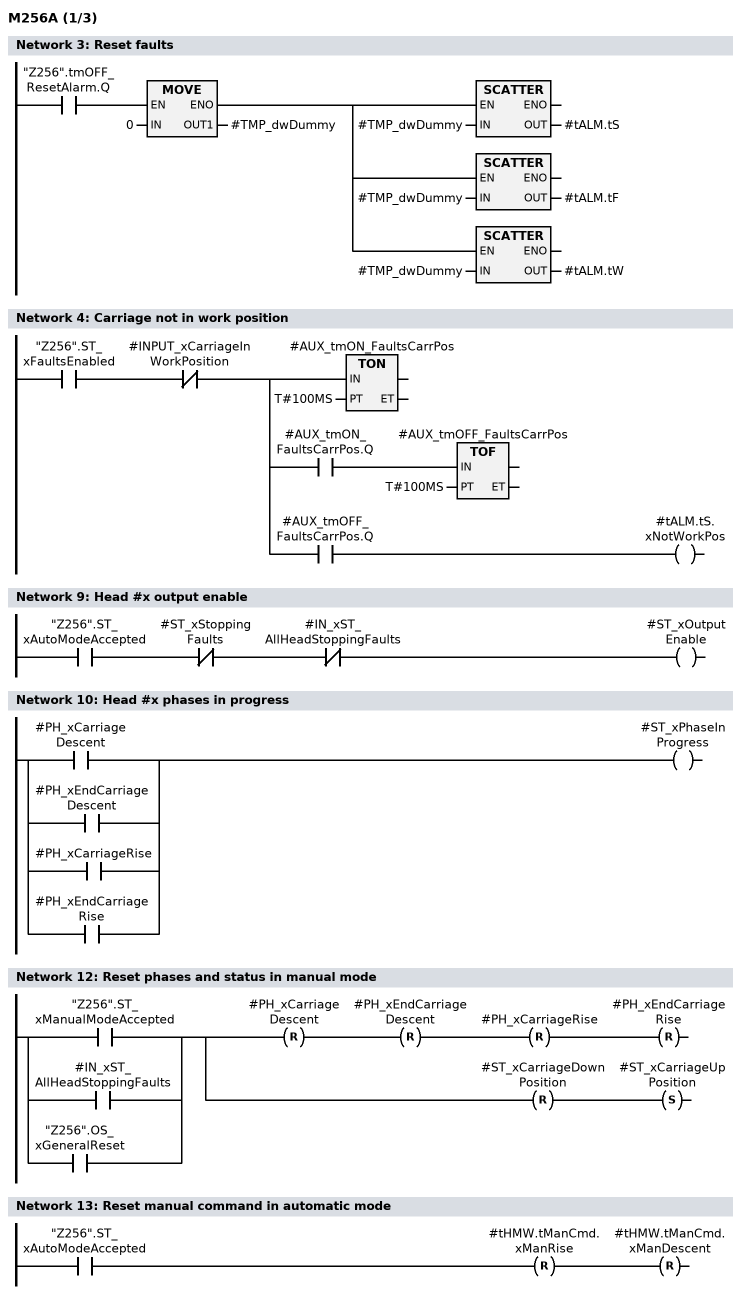
   IF "Z256".tmOFF_ResetAlarm.Q THEN #TMP_dwDummy := 0; END_IF;
   #_w1 := "Z256".tmOFF_ResetAlarm.Q;
   IF #_w1 THEN
       SCATTER(IN := #TMP_dwDummy, OUT => #tALM.tS);
       SCATTER(IN := #TMP_dwDummy, OUT => #tALM.tF);
       SCATTER(IN := #TMP_dwDummy, OUT => #tALM.tW);
   END_IF;
END_REGION

REGION Network 4: Carriage not in work position
   #_w1 := "Z256".ST_xFaultsEnabled AND NOT #INPUT_xCarriageInWorkPosition;
   #AUX_tmON_FaultsCarrPos.TON(IN := #_w1, PT := T#100MS);
   #AUX_tmOFF_FaultsCarrPos.TOF(IN := #_w1 AND #AUX_tmON_FaultsCarrPos.Q, PT := T#100MS);
   #tALM.tS.xNotWorkPos := #_w1 AND #AUX_tmOFF_FaultsCarrPos.Q;
END_REGION

REGION Network 5 (SCL): Cumulative of warning active
   #ST_xWarnings := 0;

   GATHER(IN:= #tALM.tW,
          OUT=>#TMP_dwDummy);

   IF #TMP_dwDummy <> 0 THEN
       #ST_xWarnings := 1;
   END_IF;
END_REGION

REGION Network 6 (SCL): Cumulative of stopping faults active
   #ST_xStoppingFaults := 0;
   GATHER(IN := #tALM.tS,
          OUT => #TMP_dwDummy);

   IF #TMP_dwDummy <> 0 THEN
       #ST_xStoppingFaults := 1;
   END_IF;
END_REGION

REGION Network 7 (SCL): Cumulative of faults active
   #ST_xFaults := 0;
   GATHER(IN := #tALM.tF,
          OUT => #TMP_dwDummy);

   IF #TMP_dwDummy <> 0 THEN
       #ST_xFaults := 1;
   END_IF;
END_REGION

REGION Network 8: ####_STATUS_####
END_REGION

REGION Network 9: Head #x output enable
   RUNG wire#powerrail
      Contact( "Z256".ST_xAutoModeAccepted )
      I_Contact( #ST_xStoppingFaults )
      I_Contact( #IN_xST_AllHeadStoppingFaults )
      Coil( #ST_xOutputEnable )
   END_RUNG
   // the same network as SCL:
   #ST_xOutputEnable := "Z256".ST_xAutoModeAccepted AND NOT #ST_xStoppingFaults AND NOT #IN_xST_AllHeadStoppingFaults;
END_REGION

REGION Network 10: Head #x phases in progress
   RUNG wire#powerrail
      Contact( #PH_xCarriageDescent )
      wire#w1
      Coil( #ST_xPhaseInProgress )
   END_RUNG
   RUNG wire#powerrail
      Contact( #PH_xEndCarriageDescent )
   END_RUNG wire#w1
   RUNG wire#powerrail
      Contact( #PH_xCarriageRise )
   END_RUNG wire#w1
   RUNG wire#powerrail
      Contact( #PH_xEndCarriageRise )
   END_RUNG wire#w1
   // the same network as SCL:
   #ST_xPhaseInProgress := #PH_xCarriageDescent OR #PH_xEndCarriageDescent OR #PH_xCarriageRise OR #PH_xEndCarriageRise;
END_REGION

REGION Network 11: #####_PHASES_&_LOGICS_#####
END_REGION

REGION Network 12: Reset phases and status in manual mode
   RUNG wire#powerrail
      Contact( "Z256".ST_xManualModeAccepted )
      wire#w1
      R_Coil( #PH_xCarriageDescent )
      R_Coil( #PH_xEndCarriageDescent )
      R_Coil( #PH_xCarriageRise )
      R_Coil( #PH_xEndCarriageRise )
   END_RUNG
   RUNG wire#powerrail
      Contact( #IN_xST_AllHeadStoppingFaults )
   END_RUNG wire#w1
   RUNG wire#powerrail
      Contact( "Z256".OS_xGeneralReset )
   END_RUNG wire#w1
   RUNG wire#w1
      R_Coil( #ST_xCarriageDownPosition )
      S_Coil( #ST_xCarriageUpPosition )
   END_RUNG
   // the same network as SCL:
   IF "Z256".ST_xManualModeAccepted OR #IN_xST_AllHeadStoppingFaults OR "Z256".OS_xGeneralReset THEN
       #PH_xCarriageDescent := FALSE;
       #PH_xEndCarriageDescent := FALSE;
       #PH_xCarriageRise := FALSE;
       #PH_xEndCarriageRise := FALSE;
       #ST_xCarriageDownPosition := FALSE;
       #ST_xCarriageUpPosition := TRUE;
   END_IF;
END_REGION

REGION Network 13: Reset manual command in automatic mode
   RUNG wire#powerrail
      Contact( "Z256".ST_xAutoModeAccepted )
      R_Coil( #tHMW.tManCmd.xManRise )
      R_Coil( #tHMW.tManCmd.xManDescent )
   END_RUNG
   // the same network as SCL:
   IF "Z256".ST_xAutoModeAccepted THEN
       #tHMW.tManCmd.xManRise := FALSE;
       #tHMW.tManCmd.xManDescent := FALSE;
   END_IF;
END_REGION

REGION Network 14: Carriage descent request
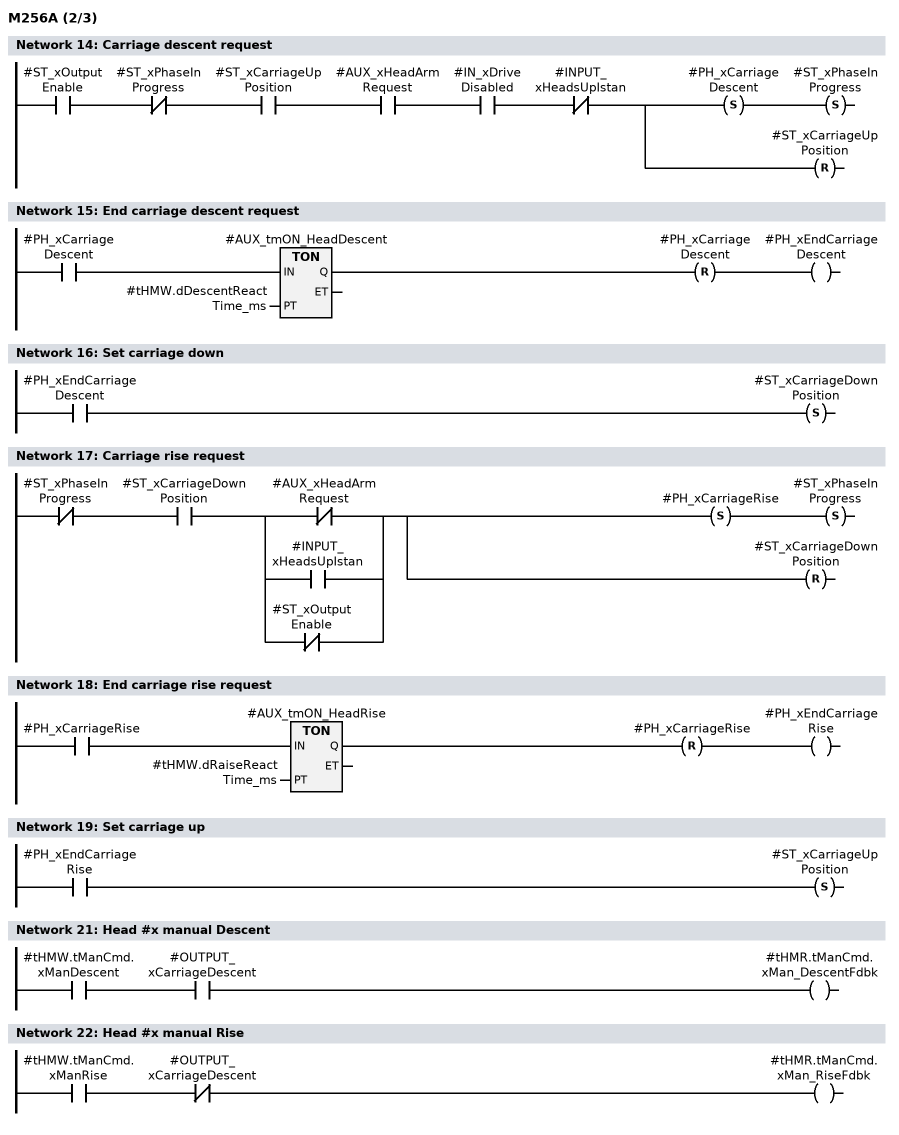
   RUNG wire#powerrail
      Contact( #ST_xOutputEnable )
      I_Contact( #ST_xPhaseInProgress )
      Contact( #ST_xCarriageUpPosition )
      Contact( #AUX_xHeadArmRequest )
      Contact( #IN_xDriveDisabled )
      I_Contact( #INPUT_xHeadsUpIstan )
      wire#w1
      S_Coil( #PH_xCarriageDescent )
      S_Coil( #ST_xPhaseInProgress )
   END_RUNG
   RUNG wire#w1
      R_Coil( #ST_xCarriageUpPosition )
   END_RUNG
   // the same network as SCL:
   IF #ST_xOutputEnable AND NOT #ST_xPhaseInProgress AND #ST_xCarriageUpPosition AND #AUX_xHeadArmRequest AND #IN_xDriveDisabled AND NOT #INPUT_xHeadsUpIstan THEN
       #PH_xCarriageDescent := TRUE;
   END_IF;
   #_w1 := #ST_xOutputEnable AND NOT #ST_xPhaseInProgress AND #ST_xCarriageUpPosition AND #AUX_xHeadArmRequest AND #IN_xDriveDisabled AND NOT #INPUT_xHeadsUpIstan;
   IF #_w1 THEN
       #ST_xPhaseInProgress := TRUE;
       #ST_xCarriageUpPosition := FALSE;
   END_IF;
END_REGION

REGION Network 15: End carriage descent request
   #AUX_tmON_HeadDescent.TON(IN := #PH_xCarriageDescent, PT := #tHMW.dDescentReactTime_ms);
   IF #AUX_tmON_HeadDescent.Q THEN #PH_xCarriageDescent := FALSE; END_IF;
   #PH_xEndCarriageDescent := #AUX_tmON_HeadDescent.Q;
END_REGION

REGION Network 16: Set carriage down
   RUNG wire#powerrail
      Contact( #PH_xEndCarriageDescent )
      S_Coil( #ST_xCarriageDownPosition )
   END_RUNG
   // the same network as SCL:
   IF #PH_xEndCarriageDescent THEN #ST_xCarriageDownPosition := TRUE; END_IF;
END_REGION

REGION Network 17: Carriage rise request
   RUNG wire#powerrail
      I_Contact( #ST_xPhaseInProgress )
      Contact( #ST_xCarriageDownPosition )
      wire#w1
      I_Contact( #AUX_xHeadArmRequest )
      wire#w2
      S_Coil( #PH_xCarriageRise )
      S_Coil( #ST_xPhaseInProgress )
   END_RUNG
   RUNG wire#w1
      Contact( #INPUT_xHeadsUpIstan )
   END_RUNG wire#w2
   RUNG wire#w1
      I_Contact( #ST_xOutputEnable )
   END_RUNG wire#w2
   RUNG wire#w2
      R_Coil( #ST_xCarriageDownPosition )
   END_RUNG
   // the same network as SCL:
   IF NOT #ST_xPhaseInProgress AND #ST_xCarriageDownPosition AND (NOT #AUX_xHeadArmRequest OR #INPUT_xHeadsUpIstan OR NOT #ST_xOutputEnable) THEN
       #PH_xCarriageRise := TRUE;
   END_IF;
   #_w1 := NOT #ST_xPhaseInProgress AND #ST_xCarriageDownPosition AND (NOT #AUX_xHeadArmRequest OR #INPUT_xHeadsUpIstan OR NOT #ST_xOutputEnable);
   IF #_w1 THEN
       #ST_xPhaseInProgress := TRUE;
       #ST_xCarriageDownPosition := FALSE;
   END_IF;
END_REGION

REGION Network 18: End carriage rise request
   #AUX_tmON_HeadRise.TON(IN := #PH_xCarriageRise, PT := #tHMW.dRaiseReactTime_ms);
   IF #AUX_tmON_HeadRise.Q THEN #PH_xCarriageRise := FALSE; END_IF;
   #PH_xEndCarriageRise := #AUX_tmON_HeadRise.Q;
END_REGION

REGION Network 19: Set carriage up
   RUNG wire#powerrail
      Contact( #PH_xEndCarriageRise )
      S_Coil( #ST_xCarriageUpPosition )
   END_RUNG
   // the same network as SCL:
   IF #PH_xEndCarriageRise THEN #ST_xCarriageUpPosition := TRUE; END_IF;
END_REGION

REGION Network 20: ### HMI STATUS ###
END_REGION

REGION Network 21: Head #x manual Descent
   RUNG wire#powerrail
      Contact( #tHMW.tManCmd.xManDescent )
      Contact( #OUTPUT_xCarriageDescent )
      Coil( #tHMR.tManCmd.xMan_DescentFdbk )
   END_RUNG
   // the same network as SCL:
   #tHMR.tManCmd.xMan_DescentFdbk := #tHMW.tManCmd.xManDescent AND #OUTPUT_xCarriageDescent;
END_REGION

REGION Network 22: Head #x manual Rise
   RUNG wire#powerrail
      Contact( #tHMW.tManCmd.xManRise )
      I_Contact( #OUTPUT_xCarriageDescent )
      Coil( #tHMR.tManCmd.xMan_RiseFdbk )
   END_RUNG
   // the same network as SCL:
   #tHMR.tManCmd.xMan_RiseFdbk := #tHMW.tManCmd.xManRise AND NOT #OUTPUT_xCarriageDescent;
END_REGION

REGION Network 23: Arm status
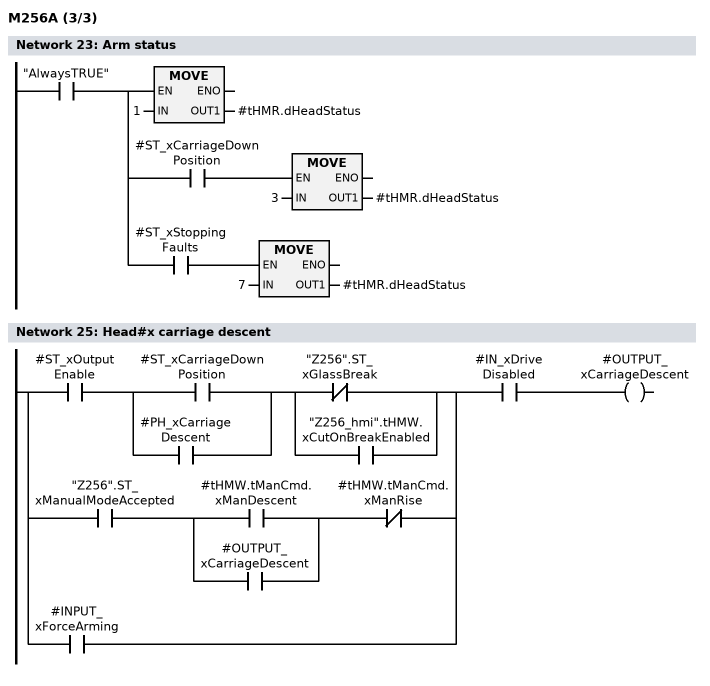
   RUNG wire#powerrail
      Contact( "AlwaysTRUE" )
      wire#w1
      Move(in := 1, out1 => #tHMR.dHeadStatus)
   END_RUNG
   RUNG wire#w1
      Contact( #ST_xCarriageDownPosition )
      Move(in := 3, out1 => #tHMR.dHeadStatus)
   END_RUNG
   RUNG wire#w1
      Contact( #ST_xStoppingFaults )
      Move(in := 7, out1 => #tHMR.dHeadStatus)
   END_RUNG
   // the same network as SCL:
   IF "AlwaysTRUE" THEN #tHMR.dHeadStatus := 1; END_IF;
   IF "AlwaysTRUE" AND #ST_xCarriageDownPosition THEN #tHMR.dHeadStatus := 3; END_IF;
   IF "AlwaysTRUE" AND #ST_xStoppingFaults THEN #tHMR.dHeadStatus := 7; END_IF;
END_REGION

REGION Network 24: ####_OUTPUT_####
END_REGION

REGION Network 25: Head#x carriage descent
   RUNG wire#powerrail
      Contact( #ST_xOutputEnable )
      wire#w1
      Contact( #ST_xCarriageDownPosition )
      wire#w2
      I_Contact( "Z256".ST_xGlassBreak )
      wire#w3
      Contact( #IN_xDriveDisabled )
      Coil( #OUTPUT_xCarriageDescent )
   END_RUNG
   RUNG wire#w1
      Contact( #PH_xCarriageDescent )
   END_RUNG wire#w2
   RUNG wire#w2
      Contact( "Z256_hmi".tHMW.xCutOnBreakEnabled )
   END_RUNG wire#w3
   RUNG wire#powerrail
      Contact( "Z256".ST_xManualModeAccepted )
      wire#w4
      Contact( #tHMW.tManCmd.xManDescent )
      wire#w5
      I_Contact( #tHMW.tManCmd.xManRise )
   END_RUNG wire#w3
   RUNG wire#w4
      Contact( #OUTPUT_xCarriageDescent )
   END_RUNG wire#w5
   RUNG wire#powerrail
      Contact( #INPUT_xForceArming )
   END_RUNG wire#w3
   // the same network as SCL:
   #OUTPUT_xCarriageDescent := ((#ST_xOutputEnable AND (#ST_xCarriageDownPosition OR #PH_xCarriageDescent) AND (NOT "Z256".ST_xGlassBreak OR "Z256_hmi".tHMW.xCutOnBreakEnabled)) OR ("Z256".ST_xManualModeAccepted AND (#tHMW.tManCmd.xManDescent OR #OUTPUT_xCarriageDescent) AND NOT #tHMW.tManCmd.xManRise) OR #INPUT_xForceArming) AND #IN_xDriveDisabled;
END_REGION
END_FUNCTION_BLOCK

FUNCTION_BLOCK "M256F"   // FB13, LAD
{ S7_Optimized_Access := 'TRUE' }
VERSION : 0.1
   VAR_INPUT
      IN_xHeadDescent : Bool;   // Head #x carriage descent
      IN_dHeadCycleIndex : DInt;   // Number of head cycle (Actual head-1)
      IN_xST_AllHeadStoppingFaults : Bool;   // Cumulative head alarm
   END_VAR
   VAR
      ST_xOutputEnable : Bool;   // Head #x output enable
      ST_xPhaseInProgress : Bool;   // Head #x phases in progress
      ST_xStoppingFaults : Bool;   // Head #x in stopping fault
      ST_xWarnings : Bool;   // Head #x in warning
      ST_xFaults : Bool;   // Head #x in faults
      OS_xPressureInc : Bool;   // OS Head #x pressure increment
      OS_xPressureDec : Bool;   // OS Head #x pressure decrement
      OSR_xPressureInc : Bool;   // OSR Head #x pressure increment
      OSR_xPressureDec : Bool;   // OSR Head #x pressure decrement
      OSR_xManEnable : Bool;   // OSR Head #x manual mode
      AUX_xFiringONRequest : Bool;   // Head #x firing ON request
      AUX_dLastCounter : DInt;   // Head #x last counter value
      AUX_dHeadUsage : DInt;   // Head #x usage mm
      AUX_xOilONRequest : Bool;   // Head #x oil ON request
      AUX_tmON_PressureInc : IEC_TIMER;   // Head #x timer ON pressure increment
      AUX_tmON_PressureDec : IEC_TIMER;   // Head #x timer ON pressure decrement
      AUX_dHeadMissionIDinProg : DInt;   // Head #x mission ID in progress
      AUX_xHeadFiringMissionInProgress : Bool;   // Head #x firing mission in progress
      OUTPUT_xFireON : Bool;   // Head #x firing ON
      OUTPUT_iPressuremA : Int;   // Head #x pressure [mA]
      OUTPUT_xOilON : Bool;   // Head #x oil ON
      INPUT_xForceFiring : Bool;   // SA Head #x firing
      INPUT_xPressureInc : Bool;   // SB Head #x pressure increment
      INPUT_xPressureDec : Bool;   // SB Head #x pressure decrement
   END_VAR
   VAR RETAIN
      tHMR : Struct   // {[Unit][Scada unit][Low limit][High limit][Access]}
         rHeadUsage_km : Real;   // Head#x head usage [km] {km|km|x|x|O}
         dHeadStatus : DInt;   // Head#x firing status (1=OFF 3=ON) {x|x|x|x|O}
         tManCmd : Struct
            xMan_FireON_Fdbk : Bool;   // Head#x manual fire ON Feeback {x|x|x|x|O}
            xMan_FireOFF_Fdbk : Bool;   // Head#x manual fire OFF Feedback {x|x|x|x|O}
            xMan_OilON_Fdbk : Bool;   // Head#x manual oil feedback ON {x|x|x|x|O}
         END_STRUCT;
      END_STRUCT;
      tHMW : Struct   // {[Unit][Scada unit][Low limit][High limit][Access]}
         dHeadFireONReaction_ms : DInt;   // Head#x fire ON reaction time [ms] {ms|s|0|1|M}
         dHeadFireOFFReaction_ms : DInt;   // Head#x fire OFF reaction time [ms] {ms|s|0|1|M}
         dHeadOilONDelay_ms : DInt;   // Head#x Oil ON delay [ms]{ms|s|-2|2|O}
         dHeadOilOFFDelay_ms : DInt;   // Head#x Oil OFF delay [ms]{ms|s|-2|2|O}
         dHeadFireONDelay_cmm : DInt;   // Head#x fire ON delay [mm/100] {mm/100|mm|-50|50|O}
         dHeadFireOFFDelay_cmm : DInt;   // Head#x fire OFF delay [mm/100] {mm/100|mm|-50|50|O}
         dHeadPressure_mN : DInt;   // Head#x pressure value [N/1000] {N/1000|N|16|180|O}
         xResetUsageCounter : Bool;   // Head#x reset head usage counter {x|x|x|x|O}
         tManCmd : Struct
            xMan_FireON : Bool;   // Head#x manual fire ON {x|x|x|x|O}
            xMan_FireOFF : Bool;   // Head#x manual fire OFF {x|x|x|x|O}
            xMan_OilON : Bool;   // Head#x manual oil ON {x|x|x|x|O}
         END_STRUCT;
      END_STRUCT;
   END_VAR
   VAR
      tALM : Struct
         tW : Struct
            x0 : Bool;
            x1 : Bool;
            x2 : Bool;
            x3 : Bool;
            x4 : Bool;
            x5 : Bool;
            x6 : Bool;
            x7 : Bool;
            x8 : Bool;
            x9 : Bool;
            x10 : Bool;
            x11 : Bool;
            x12 : Bool;
            x13 : Bool;
            x14 : Bool;
            x15 : Bool;
            x16 : Bool;
            x17 : Bool;
            x18 : Bool;
            x19 : Bool;
            x20 : Bool;
            x21 : Bool;
            x22 : Bool;
            x23 : Bool;
            x24 : Bool;
            x25 : Bool;
            x26 : Bool;
            x27 : Bool;
            x28 : Bool;
            x29 : Bool;
            x30 : Bool;
            x31 : Bool;
         END_STRUCT;
         tS : Struct
            x0 : Bool;
            x1 : Bool;
            x2 : Bool;
            x3 : Bool;
            x4 : Bool;
            x5 : Bool;
            x6 : Bool;
            x7 : Bool;
            x8 : Bool;
            x9 : Bool;
            x10 : Bool;
            x11 : Bool;
            x12 : Bool;
            x13 : Bool;
            x14 : Bool;
            x15 : Bool;
            x16 : Bool;
            x17 : Bool;
            x18 : Bool;
            x19 : Bool;
            x20 : Bool;
            x21 : Bool;
            x22 : Bool;
            x23 : Bool;
            x24 : Bool;
            x25 : Bool;
            x26 : Bool;
            x27 : Bool;
            x28 : Bool;
            x29 : Bool;
            x30 : Bool;
            x31 : Bool;
         END_STRUCT;
         tF : Struct
            x0 : Bool;
            x1 : Bool;
            x2 : Bool;
            x3 : Bool;
            x4 : Bool;
            x5 : Bool;
            x6 : Bool;
            x7 : Bool;
            x8 : Bool;
            x9 : Bool;
            x10 : Bool;
            x11 : Bool;
            x12 : Bool;
            x13 : Bool;
            x14 : Bool;
            x15 : Bool;
            x16 : Bool;
            x17 : Bool;
            x18 : Bool;
            x19 : Bool;
            x20 : Bool;
            x21 : Bool;
            x22 : Bool;
            x23 : Bool;
            x24 : Bool;
            x25 : Bool;
            x26 : Bool;
            x27 : Bool;
            x28 : Bool;
            x29 : Bool;
            x30 : Bool;
            x31 : Bool;
         END_STRUCT;
      END_STRUCT;
   END_VAR
   VAR_TEMP
      TMP_dwDummy : DWord;
      TMP_dDummy : DInt;
      TMP_rDummy : Real;
   END_VAR
   VAR_TEMP   // added for the SCL form of the ladder/FBD networks
      _w1 : Bool;
   END_VAR
BEGIN

REGION Network 1: ####_COSTANTS_####
END_REGION

REGION Network 2: ####_ALARMS_####
END_REGION

REGION Network 3: Reset faults
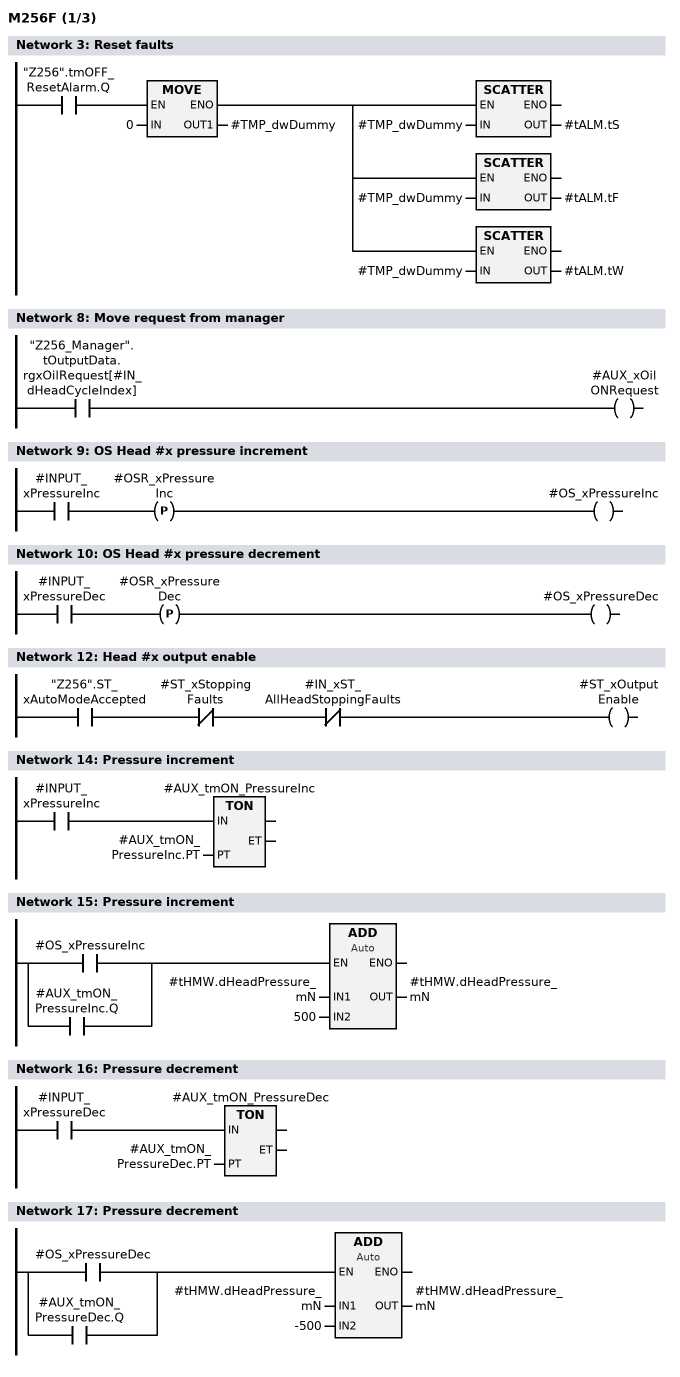
   IF "Z256".tmOFF_ResetAlarm.Q THEN #TMP_dwDummy := 0; END_IF;
   #_w1 := "Z256".tmOFF_ResetAlarm.Q;
   IF #_w1 THEN
       SCATTER(IN := #TMP_dwDummy, OUT => #tALM.tS);
       SCATTER(IN := #TMP_dwDummy, OUT => #tALM.tF);
       SCATTER(IN := #TMP_dwDummy, OUT => #tALM.tW);
   END_IF;
END_REGION

REGION Network 4 (SCL): Cumulative of warning active
   #ST_xWarnings := 0;

   GATHER(IN:= #tALM.tW,
          OUT=>#TMP_dwDummy);

   IF #TMP_dwDummy <> 0 THEN
       #ST_xWarnings := 1;
   END_IF;
END_REGION

REGION Network 5 (SCL): Cumulative of stopping faults active
   #ST_xStoppingFaults := 0;
   GATHER(IN := #tALM.tS,
          OUT => #TMP_dwDummy);

   IF #TMP_dwDummy <> 0 THEN
       #ST_xStoppingFaults := 1;
   END_IF;
END_REGION

REGION Network 6 (SCL): Cumulative of faults active
   #ST_xFaults := 0;
   GATHER(IN := #tALM.tF,
          OUT => #TMP_dwDummy);

   IF #TMP_dwDummy <> 0 THEN
       #ST_xFaults := 1;
   END_IF;
END_REGION

REGION Network 7: #####_MATCH_#####
END_REGION

REGION Network 8: Move request from manager
   RUNG wire#powerrail
      Contact( "Z256_Manager".tOutputData.rgxOilRequest[#IN_dHeadCycleIndex] )
      Coil( #AUX_xOilONRequest )
   END_RUNG
   // the same network as SCL:
   #AUX_xOilONRequest := "Z256_Manager".tOutputData.rgxOilRequest[#IN_dHeadCycleIndex];
END_REGION

REGION Network 9: OS Head #x pressure increment
   RUNG wire#powerrail
      Contact( #INPUT_xPressureInc )
      P_Trig( #OSR_xPressureInc )
      Coil( #OS_xPressureInc )
   END_RUNG
   // the same network as SCL:
   #_w1 := #INPUT_xPressureInc AND NOT #OSR_xPressureInc;   // rising edge
   #OSR_xPressureInc := #INPUT_xPressureInc;
   #OS_xPressureInc := #_w1;
END_REGION

REGION Network 10: OS Head #x pressure decrement
   RUNG wire#powerrail
      Contact( #INPUT_xPressureDec )
      P_Trig( #OSR_xPressureDec )
      Coil( #OS_xPressureDec )
   END_RUNG
   // the same network as SCL:
   #_w1 := #INPUT_xPressureDec AND NOT #OSR_xPressureDec;   // rising edge
   #OSR_xPressureDec := #INPUT_xPressureDec;
   #OS_xPressureDec := #_w1;
END_REGION

REGION Network 11: #####_STATUSES_#####
END_REGION

REGION Network 12: Head #x output enable
   RUNG wire#powerrail
      Contact( "Z256".ST_xAutoModeAccepted )
      I_Contact( #ST_xStoppingFaults )
      I_Contact( #IN_xST_AllHeadStoppingFaults )
      Coil( #ST_xOutputEnable )
   END_RUNG
   // the same network as SCL:
   #ST_xOutputEnable := "Z256".ST_xAutoModeAccepted AND NOT #ST_xStoppingFaults AND NOT #IN_xST_AllHeadStoppingFaults;
END_REGION

REGION Network 13: #####_PHASES&LOGICS_#####
END_REGION

REGION Network 14: Pressure increment
   #AUX_tmON_PressureInc.TON(IN := #INPUT_xPressureInc, PT := #AUX_tmON_PressureInc.PT);
END_REGION

REGION Network 15: Pressure increment
   RUNG wire#powerrail
      Contact( #OS_xPressureInc )
      wire#w1
      Add(in1 := #tHMW.dHeadPressure_mN, in2 := 500, out => #tHMW.dHeadPressure_mN)
   END_RUNG
   RUNG wire#powerrail
      Contact( #AUX_tmON_PressureInc.Q )
   END_RUNG wire#w1
   // the same network as SCL:
   IF #OS_xPressureInc OR #AUX_tmON_PressureInc.Q THEN
       #tHMW.dHeadPressure_mN := #tHMW.dHeadPressure_mN + 500;
   END_IF;
END_REGION

REGION Network 16: Pressure decrement
   #AUX_tmON_PressureDec.TON(IN := #INPUT_xPressureDec, PT := #AUX_tmON_PressureDec.PT);
END_REGION

REGION Network 17: Pressure decrement
   RUNG wire#powerrail
      Contact( #OS_xPressureDec )
      wire#w1
      Add(in1 := #tHMW.dHeadPressure_mN, in2 := -500, out => #tHMW.dHeadPressure_mN)
   END_RUNG
   RUNG wire#powerrail
      Contact( #AUX_tmON_PressureDec.Q )
   END_RUNG wire#w1
   // the same network as SCL:
   IF #OS_xPressureDec OR #AUX_tmON_PressureDec.Q THEN
       #tHMW.dHeadPressure_mN := #tHMW.dHeadPressure_mN + (-500);
   END_IF;
END_REGION

REGION Network 18: Check pressure imits
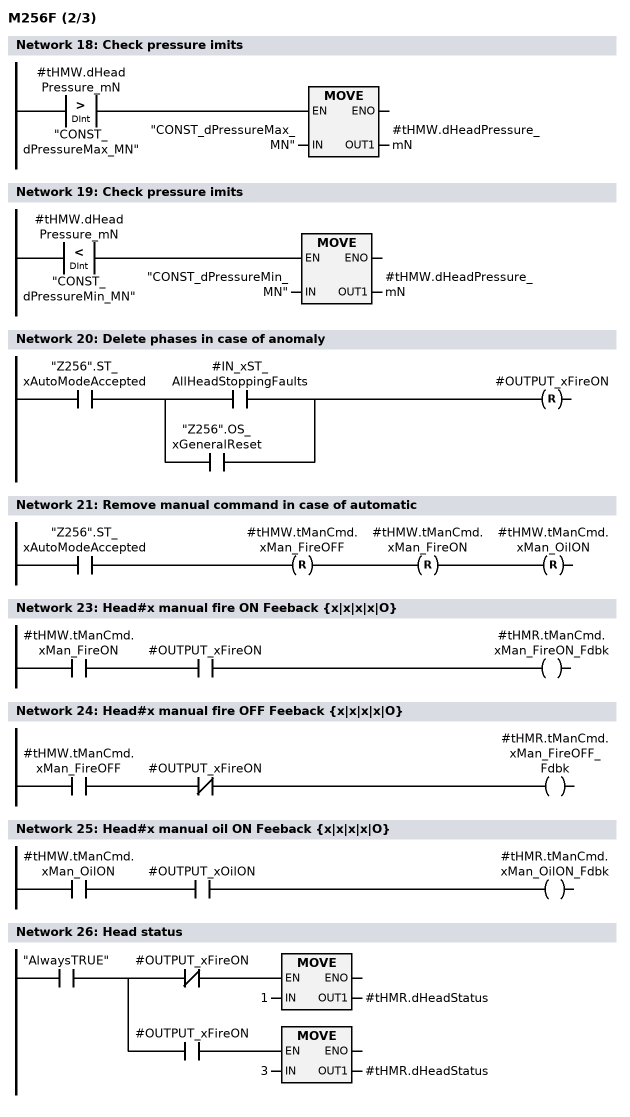
   RUNG wire#powerrail
      { S7_Templates := "SrcType := DInt" } GT_Contact(in1 := #tHMW.dHeadPressure_mN, in2 := "CONST_dPressureMax_MN")
      Move(in := "CONST_dPressureMax_MN", out1 => #tHMW.dHeadPressure_mN)
   END_RUNG
   // the same network as SCL:
   IF #tHMW.dHeadPressure_mN > "CONST_dPressureMax_MN" THEN
       #tHMW.dHeadPressure_mN := "CONST_dPressureMax_MN";
   END_IF;
END_REGION

REGION Network 19: Check pressure imits
   RUNG wire#powerrail
      { S7_Templates := "SrcType := DInt" } LT_Contact(in1 := #tHMW.dHeadPressure_mN, in2 := "CONST_dPressureMin_MN")
      Move(in := "CONST_dPressureMin_MN", out1 => #tHMW.dHeadPressure_mN)
   END_RUNG
   // the same network as SCL:
   IF #tHMW.dHeadPressure_mN < "CONST_dPressureMin_MN" THEN
       #tHMW.dHeadPressure_mN := "CONST_dPressureMin_MN";
   END_IF;
END_REGION

REGION Network 20: Delete phases in case of anomaly
   RUNG wire#powerrail
      Contact( "Z256".ST_xAutoModeAccepted )
      wire#w1
      Contact( #IN_xST_AllHeadStoppingFaults )
      wire#w2
      R_Coil( #OUTPUT_xFireON )
   END_RUNG
   RUNG wire#w1
      Contact( "Z256".OS_xGeneralReset )
   END_RUNG wire#w2
   // the same network as SCL:
   IF "Z256".ST_xAutoModeAccepted AND (#IN_xST_AllHeadStoppingFaults OR "Z256".OS_xGeneralReset) THEN
       #OUTPUT_xFireON := FALSE;
   END_IF;
END_REGION

REGION Network 21: Remove manual command in case of automatic
   RUNG wire#powerrail
      Contact( "Z256".ST_xAutoModeAccepted )
      R_Coil( #tHMW.tManCmd.xMan_FireOFF )
      R_Coil( #tHMW.tManCmd.xMan_FireON )
      R_Coil( #tHMW.tManCmd.xMan_OilON )
   END_RUNG
   // the same network as SCL:
   IF "Z256".ST_xAutoModeAccepted THEN
       #tHMW.tManCmd.xMan_FireOFF := FALSE;
       #tHMW.tManCmd.xMan_FireON := FALSE;
       #tHMW.tManCmd.xMan_OilON := FALSE;
   END_IF;
END_REGION

REGION Network 22: ### HMI STATUS ###
END_REGION

REGION Network 23: Head#x manual fire ON Feeback {x|x|x|x|O}
   RUNG wire#powerrail
      Contact( #tHMW.tManCmd.xMan_FireON )
      Contact( #OUTPUT_xFireON )
      Coil( #tHMR.tManCmd.xMan_FireON_Fdbk )
   END_RUNG
   // the same network as SCL:
   #tHMR.tManCmd.xMan_FireON_Fdbk := #tHMW.tManCmd.xMan_FireON AND #OUTPUT_xFireON;
END_REGION

REGION Network 24: Head#x manual fire OFF Feeback {x|x|x|x|O}
   RUNG wire#powerrail
      Contact( #tHMW.tManCmd.xMan_FireOFF )
      I_Contact( #OUTPUT_xFireON )
      Coil( #tHMR.tManCmd.xMan_FireOFF_Fdbk )
   END_RUNG
   // the same network as SCL:
   #tHMR.tManCmd.xMan_FireOFF_Fdbk := #tHMW.tManCmd.xMan_FireOFF AND NOT #OUTPUT_xFireON;
END_REGION

REGION Network 25: Head#x manual oil ON Feeback {x|x|x|x|O}
   RUNG wire#powerrail
      Contact( #tHMW.tManCmd.xMan_OilON )
      Contact( #OUTPUT_xOilON )
      Coil( #tHMR.tManCmd.xMan_OilON_Fdbk )
   END_RUNG
   // the same network as SCL:
   #tHMR.tManCmd.xMan_OilON_Fdbk := #tHMW.tManCmd.xMan_OilON AND #OUTPUT_xOilON;
END_REGION

REGION Network 26: Head status
   RUNG wire#powerrail
      Contact( "AlwaysTRUE" )
      wire#w1
      I_Contact( #OUTPUT_xFireON )
      Move(in := 1, out1 => #tHMR.dHeadStatus)
   END_RUNG
   RUNG wire#w1
      Contact( #OUTPUT_xFireON )
      Move(in := 3, out1 => #tHMR.dHeadStatus)
   END_RUNG
   // the same network as SCL:
   IF "AlwaysTRUE" AND NOT #OUTPUT_xFireON THEN #tHMR.dHeadStatus := 1; END_IF;
   IF "AlwaysTRUE" AND #OUTPUT_xFireON THEN #tHMR.dHeadStatus := 3; END_IF;
END_REGION

REGION Network 27: Head#x reset head usage counter {x|x|x|x|O}
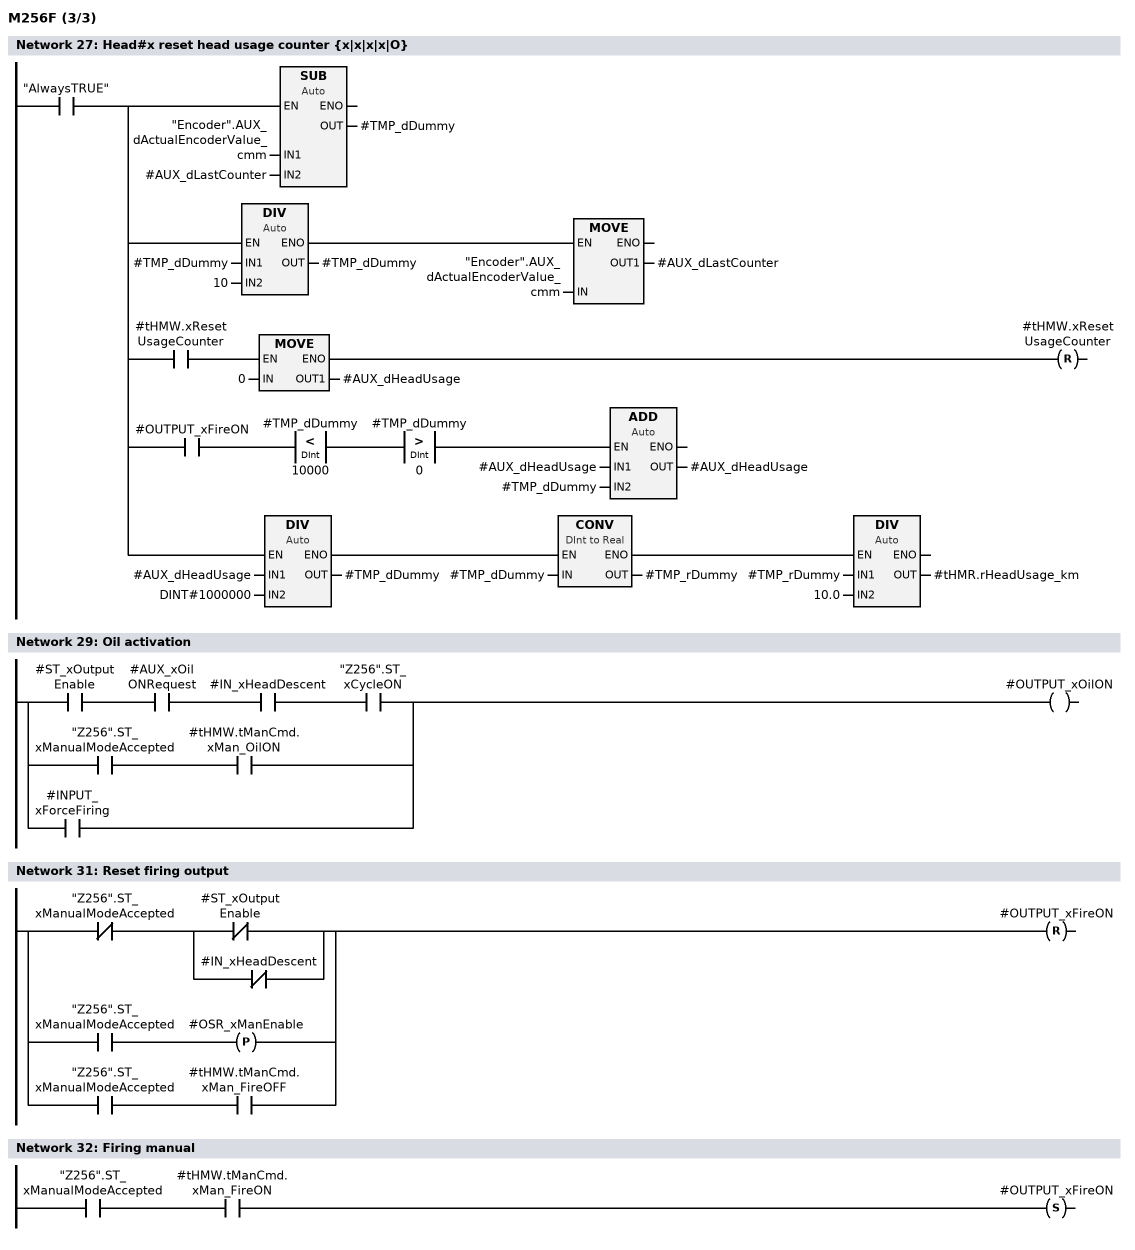
   RUNG wire#powerrail
      Contact( "AlwaysTRUE" )
      wire#w1
      Sub(in1 := "Encoder".AUX_dActualEncoderValue_cmm, in2 := #AUX_dLastCounter, out => #TMP_dDummy)
   END_RUNG
   RUNG wire#w1
      Div(in1 := #TMP_dDummy, in2 := 10, out => #TMP_dDummy)
      Move(in := "Encoder".AUX_dActualEncoderValue_cmm, out1 => #AUX_dLastCounter)
   END_RUNG
   RUNG wire#w1
      Contact( #tHMW.xResetUsageCounter )
      Move(in := 0, out1 => #AUX_dHeadUsage)
      R_Coil( #tHMW.xResetUsageCounter )
   END_RUNG
   RUNG wire#w1
      Contact( #OUTPUT_xFireON )
      { S7_Templates := "SrcType := DInt" } LT_Contact(in1 := #TMP_dDummy, in2 := 10000)
      { S7_Templates := "SrcType := DInt" } GT_Contact(in1 := #TMP_dDummy, in2 := 0)
      Add(in1 := #AUX_dHeadUsage, in2 := #TMP_dDummy, out => #AUX_dHeadUsage)
   END_RUNG
   RUNG wire#w1
      Div(in1 := #AUX_dHeadUsage, in2 := DINT#1000000, out => #TMP_dDummy)
      { S7_Templates := "[SrcType := DInt, DestType := Real]" } Convert(in := #TMP_dDummy, out => #TMP_rDummy)
      Div(in1 := #TMP_rDummy, in2 := 10.0, out => #tHMR.rHeadUsage_km)
   END_RUNG
   // the same network as SCL:
   IF "AlwaysTRUE" THEN
       #TMP_dDummy := "Encoder".AUX_dActualEncoderValue_cmm - #AUX_dLastCounter;
       #TMP_dDummy := #TMP_dDummy / 10;
       #AUX_dLastCounter := "Encoder".AUX_dActualEncoderValue_cmm;
   END_IF;
   IF "AlwaysTRUE" AND #tHMW.xResetUsageCounter THEN
       #AUX_dHeadUsage := 0;
       #tHMW.xResetUsageCounter := FALSE;
   END_IF;
   IF "AlwaysTRUE" AND #OUTPUT_xFireON AND (#TMP_dDummy < 10000) AND (#TMP_dDummy > 0) THEN
       #AUX_dHeadUsage := #AUX_dHeadUsage + #TMP_dDummy;
   END_IF;
   IF "AlwaysTRUE" THEN
       #TMP_dDummy := #AUX_dHeadUsage / DINT#1000000;
       #TMP_rDummy := DINT_TO_REAL(#TMP_dDummy);
       #tHMR.rHeadUsage_km := #TMP_rDummy / 10.0;
   END_IF;
END_REGION

REGION Network 28: ####_OUTPUT_####
END_REGION

REGION Network 29: Oil activation
   RUNG wire#powerrail
      Contact( #ST_xOutputEnable )
      Contact( #AUX_xOilONRequest )
      Contact( #IN_xHeadDescent )
      Contact( "Z256".ST_xCycleON )
      wire#w1
      Coil( #OUTPUT_xOilON )
   END_RUNG
   RUNG wire#powerrail
      Contact( "Z256".ST_xManualModeAccepted )
      Contact( #tHMW.tManCmd.xMan_OilON )
   END_RUNG wire#w1
   RUNG wire#powerrail
      Contact( #INPUT_xForceFiring )
   END_RUNG wire#w1
   // the same network as SCL:
   #OUTPUT_xOilON := (#ST_xOutputEnable AND #AUX_xOilONRequest AND #IN_xHeadDescent AND "Z256".ST_xCycleON) OR ("Z256".ST_xManualModeAccepted AND #tHMW.tManCmd.xMan_OilON) OR #INPUT_xForceFiring;
END_REGION

REGION Network 30 (SCL): Pressure to heads and display
   #TMP_rDummy := DINT_TO_REAL("CONST_dPressureMax_Unit"-"CONST_dPressureMin_Unit")/ DINT_TO_REAL("CONST_dPressureMax_MN"-"CONST_dPressureMin_MN");
   #TMP_dDummy :=#tHMW.dHeadPressure_mN-"CONST_dPressureMin_MN";
   #OUTPUT_iPressuremA := REAL_TO_INT(#TMP_rDummy *  DINT_TO_REAL(#TMP_dDummy))+DINT_TO_INT("CONST_dPressureMin_Unit");

   IF "CM_IDEV_FromMainLine".xQLTplate THEN
       #OUTPUT_iPressuremA := #OUTPUT_iPressuremA / 100 * DINT_TO_INT("Z256_hmi".tHMW.dPressureScalerOnSample_perc);
   END_IF;
END_REGION

REGION Network 31: Reset firing output
   RUNG wire#powerrail
      I_Contact( "Z256".ST_xManualModeAccepted )
      wire#w1
      I_Contact( #ST_xOutputEnable )
      wire#w2
      R_Coil( #OUTPUT_xFireON )
   END_RUNG
   RUNG wire#w1
      I_Contact( #IN_xHeadDescent )
   END_RUNG wire#w2
   RUNG wire#powerrail
      Contact( "Z256".ST_xManualModeAccepted )
      P_Trig( #OSR_xManEnable )
   END_RUNG wire#w2
   RUNG wire#powerrail
      Contact( "Z256".ST_xManualModeAccepted )
      Contact( #tHMW.tManCmd.xMan_FireOFF )
   END_RUNG wire#w2
   // the same network as SCL:
   #_w1 := "Z256".ST_xManualModeAccepted AND NOT #OSR_xManEnable;   // rising edge
   #OSR_xManEnable := "Z256".ST_xManualModeAccepted;
   IF (NOT "Z256".ST_xManualModeAccepted AND (NOT #ST_xOutputEnable OR NOT #IN_xHeadDescent)) OR #_w1 OR ("Z256".ST_xManualModeAccepted AND #tHMW.tManCmd.xMan_FireOFF) THEN
       #OUTPUT_xFireON := FALSE;
   END_IF;
END_REGION

REGION Network 32: Firing manual
   RUNG wire#powerrail
      Contact( "Z256".ST_xManualModeAccepted )
      Contact( #tHMW.tManCmd.xMan_FireON )
      S_Coil( #OUTPUT_xFireON )
   END_RUNG
   // the same network as SCL:
   IF "Z256".ST_xManualModeAccepted AND #tHMW.tManCmd.xMan_FireON THEN #OUTPUT_xFireON := TRUE; END_IF;
END_REGION
END_FUNCTION_BLOCK

FUNCTION_BLOCK "M256M"   // FB101, LAD
{ S7_Optimized_Access := 'TRUE' }